(* Logix 5000 project; controller _GigaDiscovery vendor 1 type 14 code 244 rev 35.11; software revision 35.03; part 19 of 23 *)
(* tags used below, declared in another part *)
   CROUT_Air_Compressor : UDT_CROUT;   // Compressor Command -Q18101E
   I_Platform_Closed : UDT_DCM;   // Platform Closed RFID Series -B22501J... -B22807J -B22801B
   I_Platform_Opened : UDT_DCM;   // Platform Opened RFID Series -Q23801J -Q23807J
   No_Sfty : Std_to_Sfty;
   O_Close_Platform : BOOL;
   O_Compressor_Cmd : BOOL;
   O_Open_Platform : BOOL;
   O_Pilots_Valve_Platform : BOOL;
   O_Platform_Main_Valve : BOOL;   // Valvola principale piattaforma B21902I
   O_Platform_MainValve : UDT_CROUT;   // Platform main valve B21902I
   Platform_CloseMain_Valve_Aux_Comand : BOOL;   // Valvola principale piattaforma QV6515E
   Platform_Fbk_Valv_Close : BOOL;   // Platform Close Main Valve Limit Switch -B21909I
   Platform_Fbk_Valv_Open : BOOL;   // Platform Open Main Valve Limit Switch -B21905I
   Platform_OpenMain_Valve_Aux_Comand : BOOL;   // Valvola principale piattaforma QV6515E
   Reset_Pulse : BOOL;
   RESTRAINTS_Rack : LapBar_Racks[41];
   RESTRAINTS_Sector : LapBars_Sector[9];
   Valve_Proof_Test_Cycle : Sequencer;
   Valves_Pressure_Discrepancy : DINT;
(* S_Output, continued *)

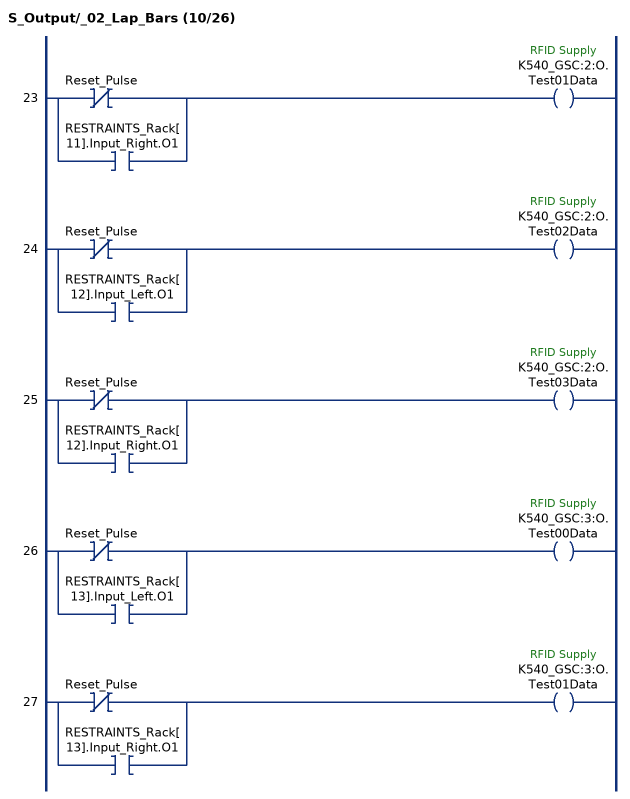
   [picture p369: S_Output/_02_Lap_Bars rungs 23-27]
   23: [XIO(Reset_Pulse) ,XIC(RESTRAINTS_Rack[11].Input_Right.O1) ]OTE(K540_GSC:2:O.Test01Data);
   24: [XIO(Reset_Pulse) ,XIC(RESTRAINTS_Rack[12].Input_Left.O1) ]OTE(K540_GSC:2:O.Test02Data);
   25: [XIO(Reset_Pulse) ,XIC(RESTRAINTS_Rack[12].Input_Right.O1) ]OTE(K540_GSC:2:O.Test03Data);
   26: [XIO(Reset_Pulse) ,XIC(RESTRAINTS_Rack[13].Input_Left.O1) ]OTE(K540_GSC:3:O.Test00Data);
   27: [XIO(Reset_Pulse) ,XIC(RESTRAINTS_Rack[13].Input_Right.O1) ]OTE(K540_GSC:3:O.Test01Data);
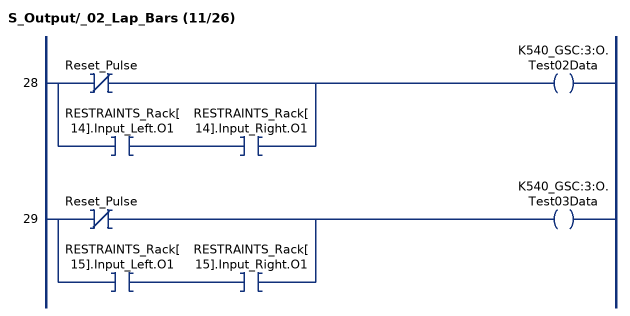
   28: [XIO(Reset_Pulse) ,XIC(RESTRAINTS_Rack[14].Input_Left.O1) XIC(RESTRAINTS_Rack[14].Input_Right.O1) ]OTE(K540_GSC:3:O.Test02Data);
   29: [XIO(Reset_Pulse) ,XIC(RESTRAINTS_Rack[15].Input_Left.O1) XIC(RESTRAINTS_Rack[15].Input_Right.O1) ]OTE(K540_GSC:3:O.Test03Data);
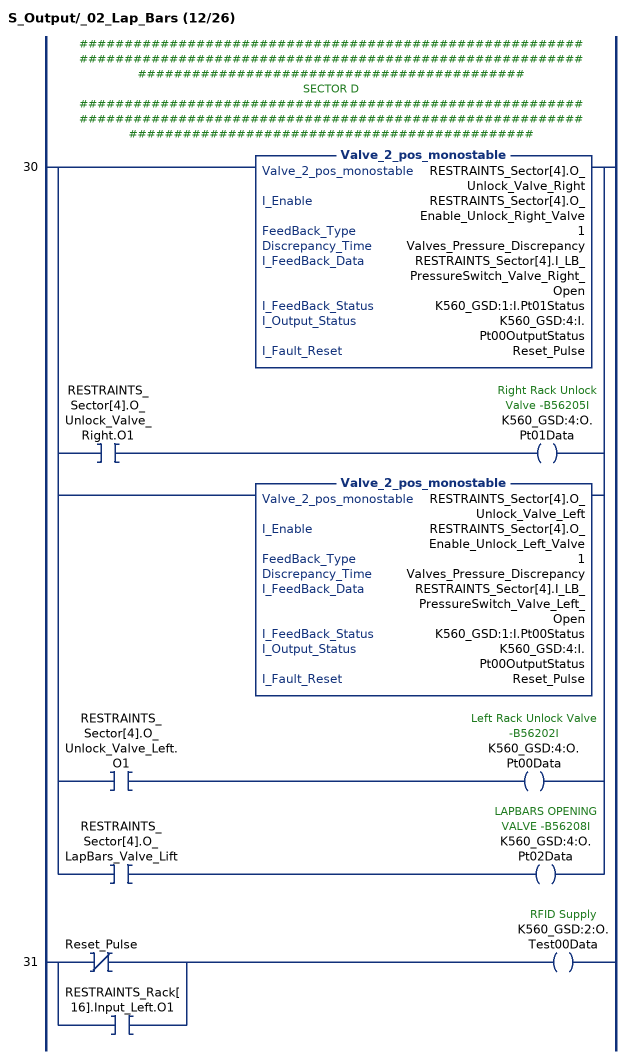
   // ###########################################################################################################################################################
   // SECTOR D
   // #############################################################################################################################################################
   30: [[Valve_2_pos_monostable(RESTRAINTS_Sector[4].O_Unlock_Valve_Right,RESTRAINTS_Sector[4].O_Enable_Unlock_Right_Valve,1,Valves_Pressure_Discrepancy,RESTRAINTS_Sector[4].I_LB_PressureSwitch_Valve_Right_Open,K560_GSD:1:I.Pt01Status,K560_GSD:4:I.Pt00OutputStatus,Reset_Pulse) ,XIC(RESTRAINTS_Sector[4].O_Unlock_Valve_Right.O1) OTE(K560_GSD:4:O.Pt01Data) ] ,[Valve_2_pos_monostable(RESTRAINTS_Sector[4].O_Unlock_Valve_Left,RESTRAINTS_Sector[4].O_Enable_Unlock_Left_Valve,1,Valves_Pressure_Discrepancy,RESTRAINTS_Sector[4].I_LB_PressureSwitch_Valve_Left_Open,K560_GSD:1:I.Pt00Status,K560_GSD:4:I.Pt00OutputStatus,Reset_Pulse) ,XIC(RESTRAINTS_Sector[4].O_Unlock_Valve_Left.O1) OTE(K560_GSD:4:O.Pt00Data) ] ,XIC(RESTRAINTS_Sector[4].O_LapBars_Valve_Lift) OTE(K560_GSD:4:O.Pt02Data) ];
   31: [XIO(Reset_Pulse) ,XIC(RESTRAINTS_Rack[16].Input_Left.O1) ]OTE(K560_GSD:2:O.Test00Data);
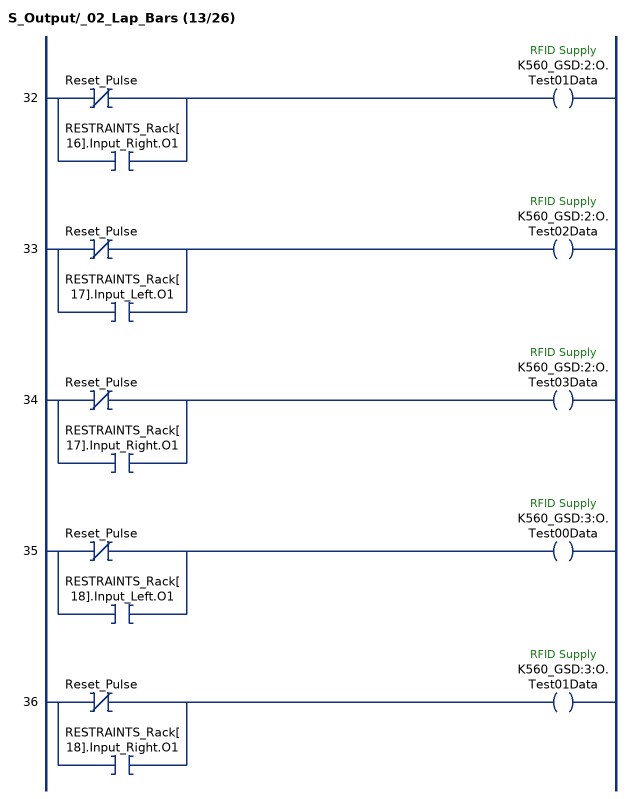
   32: [XIO(Reset_Pulse) ,XIC(RESTRAINTS_Rack[16].Input_Right.O1) ]OTE(K560_GSD:2:O.Test01Data);
   33: [XIO(Reset_Pulse) ,XIC(RESTRAINTS_Rack[17].Input_Left.O1) ]OTE(K560_GSD:2:O.Test02Data);
   34: [XIO(Reset_Pulse) ,XIC(RESTRAINTS_Rack[17].Input_Right.O1) ]OTE(K560_GSD:2:O.Test03Data);
   35: [XIO(Reset_Pulse) ,XIC(RESTRAINTS_Rack[18].Input_Left.O1) ]OTE(K560_GSD:3:O.Test00Data);
   36: [XIO(Reset_Pulse) ,XIC(RESTRAINTS_Rack[18].Input_Right.O1) ]OTE(K560_GSD:3:O.Test01Data);
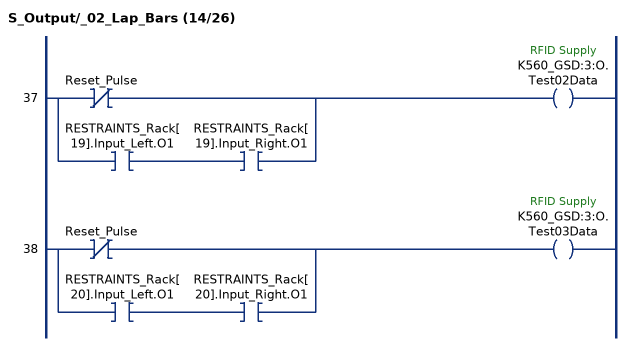
   37: [XIO(Reset_Pulse) ,XIC(RESTRAINTS_Rack[19].Input_Left.O1) XIC(RESTRAINTS_Rack[19].Input_Right.O1) ]OTE(K560_GSD:3:O.Test02Data);
   38: [XIO(Reset_Pulse) ,XIC(RESTRAINTS_Rack[20].Input_Left.O1) XIC(RESTRAINTS_Rack[20].Input_Right.O1) ]OTE(K560_GSD:3:O.Test03Data);
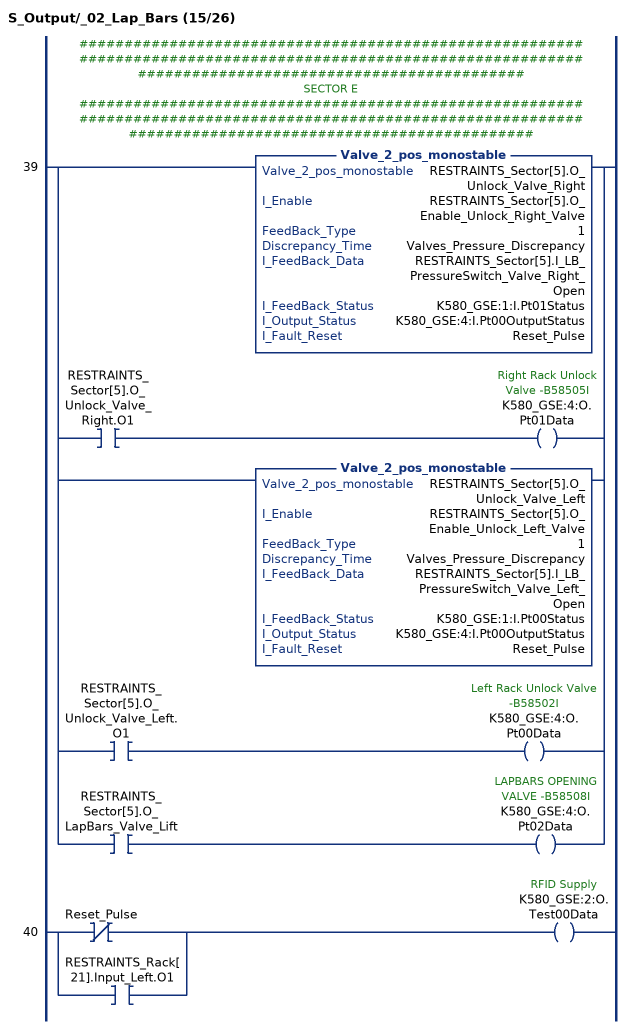
   // ###########################################################################################################################################################
   // SECTOR E
   // #############################################################################################################################################################
   39: [[Valve_2_pos_monostable(RESTRAINTS_Sector[5].O_Unlock_Valve_Right,RESTRAINTS_Sector[5].O_Enable_Unlock_Right_Valve,1,Valves_Pressure_Discrepancy,RESTRAINTS_Sector[5].I_LB_PressureSwitch_Valve_Right_Open,K580_GSE:1:I.Pt01Status,K580_GSE:4:I.Pt00OutputStatus,Reset_Pulse) ,XIC(RESTRAINTS_Sector[5].O_Unlock_Valve_Right.O1) OTE(K580_GSE:4:O.Pt01Data) ] ,[Valve_2_pos_monostable(RESTRAINTS_Sector[5].O_Unlock_Valve_Left,RESTRAINTS_Sector[5].O_Enable_Unlock_Left_Valve,1,Valves_Pressure_Discrepancy,RESTRAINTS_Sector[5].I_LB_PressureSwitch_Valve_Left_Open,K580_GSE:1:I.Pt00Status,K580_GSE:4:I.Pt00OutputStatus,Reset_Pulse) ,XIC(RESTRAINTS_Sector[5].O_Unlock_Valve_Left.O1) OTE(K580_GSE:4:O.Pt00Data) ] ,XIC(RESTRAINTS_Sector[5].O_LapBars_Valve_Lift) OTE(K580_GSE:4:O.Pt02Data) ];
   40: [XIO(Reset_Pulse) ,XIC(RESTRAINTS_Rack[21].Input_Left.O1) ]OTE(K580_GSE:2:O.Test00Data);
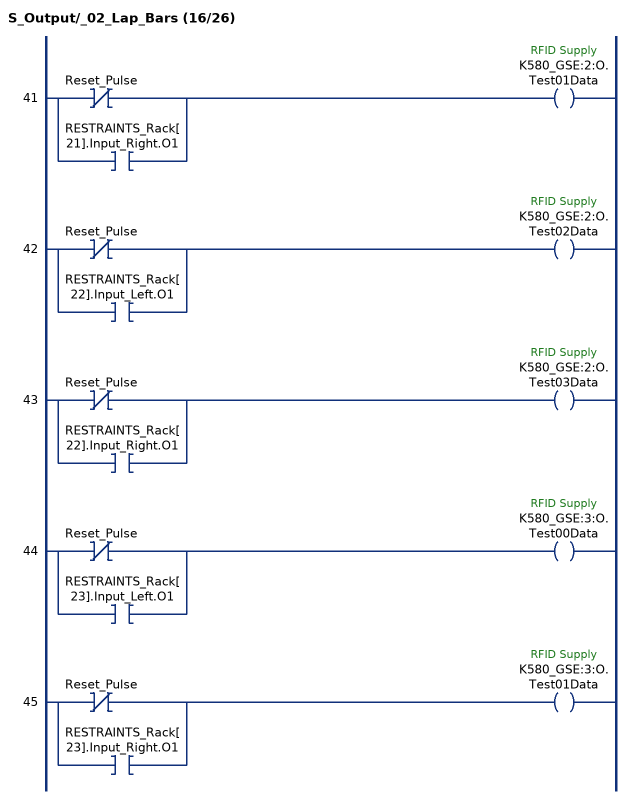
   41: [XIO(Reset_Pulse) ,XIC(RESTRAINTS_Rack[21].Input_Right.O1) ]OTE(K580_GSE:2:O.Test01Data);
   42: [XIO(Reset_Pulse) ,XIC(RESTRAINTS_Rack[22].Input_Left.O1) ]OTE(K580_GSE:2:O.Test02Data);
   43: [XIO(Reset_Pulse) ,XIC(RESTRAINTS_Rack[22].Input_Right.O1) ]OTE(K580_GSE:2:O.Test03Data);
   44: [XIO(Reset_Pulse) ,XIC(RESTRAINTS_Rack[23].Input_Left.O1) ]OTE(K580_GSE:3:O.Test00Data);
   45: [XIO(Reset_Pulse) ,XIC(RESTRAINTS_Rack[23].Input_Right.O1) ]OTE(K580_GSE:3:O.Test01Data);
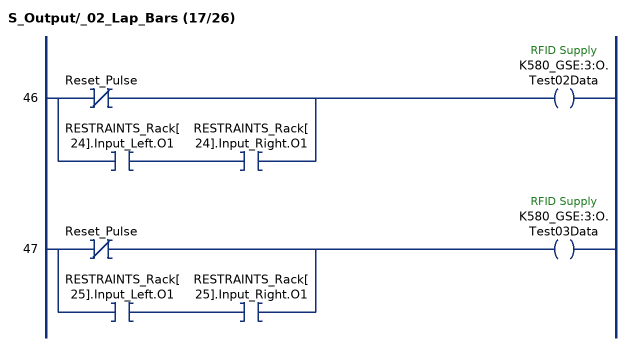
   46: [XIO(Reset_Pulse) ,XIC(RESTRAINTS_Rack[24].Input_Left.O1) XIC(RESTRAINTS_Rack[24].Input_Right.O1) ]OTE(K580_GSE:3:O.Test02Data);
   47: [XIO(Reset_Pulse) ,XIC(RESTRAINTS_Rack[25].Input_Left.O1) XIC(RESTRAINTS_Rack[25].Input_Right.O1) ]OTE(K580_GSE:3:O.Test03Data);
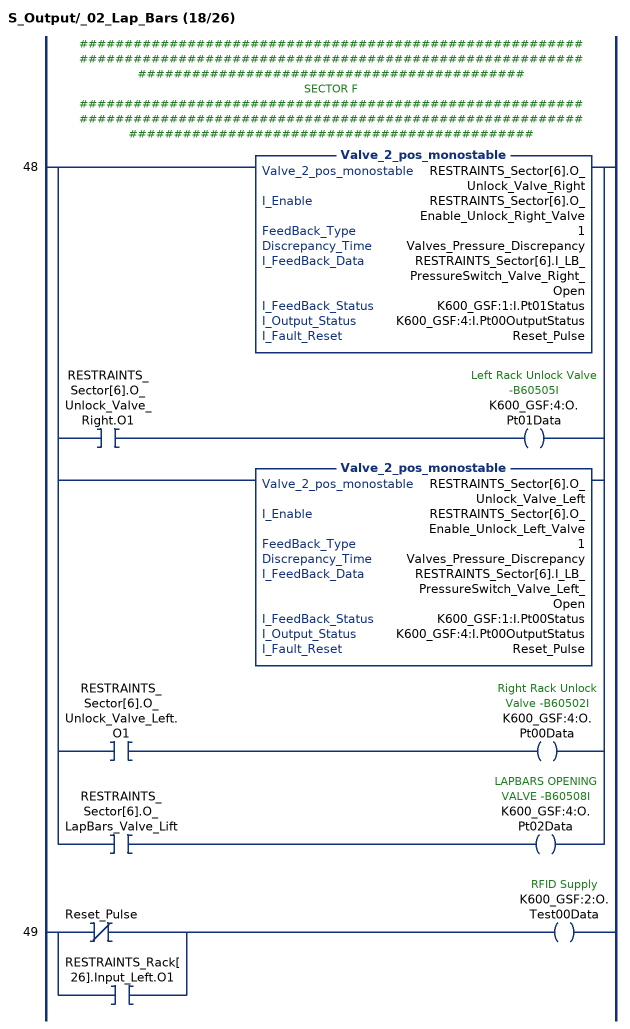
   // ###########################################################################################################################################################
   // SECTOR F
   // #############################################################################################################################################################
   48: [[Valve_2_pos_monostable(RESTRAINTS_Sector[6].O_Unlock_Valve_Right,RESTRAINTS_Sector[6].O_Enable_Unlock_Right_Valve,1,Valves_Pressure_Discrepancy,RESTRAINTS_Sector[6].I_LB_PressureSwitch_Valve_Right_Open,K600_GSF:1:I.Pt01Status,K600_GSF:4:I.Pt00OutputStatus,Reset_Pulse) ,XIC(RESTRAINTS_Sector[6].O_Unlock_Valve_Right.O1) OTE(K600_GSF:4:O.Pt01Data) ] ,[Valve_2_pos_monostable(RESTRAINTS_Sector[6].O_Unlock_Valve_Left,RESTRAINTS_Sector[6].O_Enable_Unlock_Left_Valve,1,Valves_Pressure_Discrepancy,RESTRAINTS_Sector[6].I_LB_PressureSwitch_Valve_Left_Open,K600_GSF:1:I.Pt00Status,K600_GSF:4:I.Pt00OutputStatus,Reset_Pulse) ,XIC(RESTRAINTS_Sector[6].O_Unlock_Valve_Left.O1) OTE(K600_GSF:4:O.Pt00Data) ] ,XIC(RESTRAINTS_Sector[6].O_LapBars_Valve_Lift) OTE(K600_GSF:4:O.Pt02Data) ];
   49: [XIO(Reset_Pulse) ,XIC(RESTRAINTS_Rack[26].Input_Left.O1) ]OTE(K600_GSF:2:O.Test00Data);
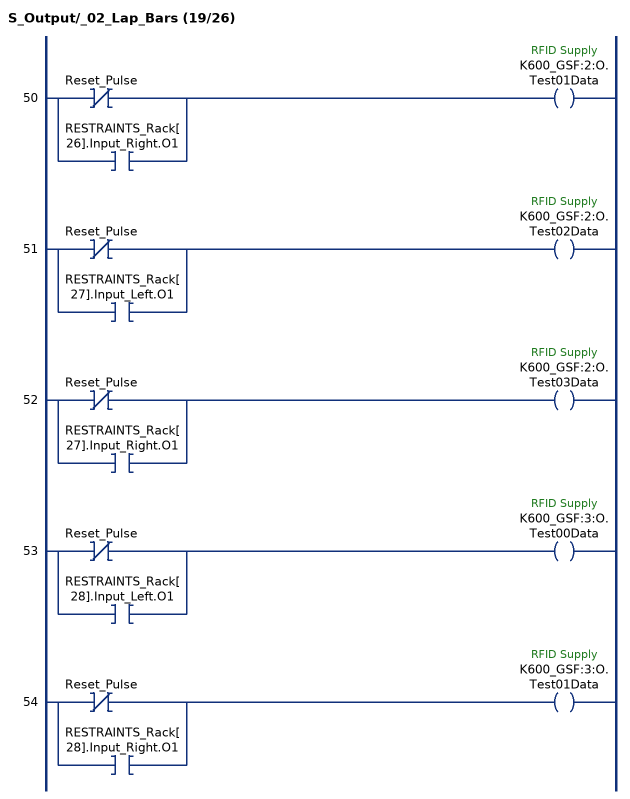
   50: [XIO(Reset_Pulse) ,XIC(RESTRAINTS_Rack[26].Input_Right.O1) ]OTE(K600_GSF:2:O.Test01Data);
   51: [XIO(Reset_Pulse) ,XIC(RESTRAINTS_Rack[27].Input_Left.O1) ]OTE(K600_GSF:2:O.Test02Data);
   52: [XIO(Reset_Pulse) ,XIC(RESTRAINTS_Rack[27].Input_Right.O1) ]OTE(K600_GSF:2:O.Test03Data);
   53: [XIO(Reset_Pulse) ,XIC(RESTRAINTS_Rack[28].Input_Left.O1) ]OTE(K600_GSF:3:O.Test00Data);
   54: [XIO(Reset_Pulse) ,XIC(RESTRAINTS_Rack[28].Input_Right.O1) ]OTE(K600_GSF:3:O.Test01Data);
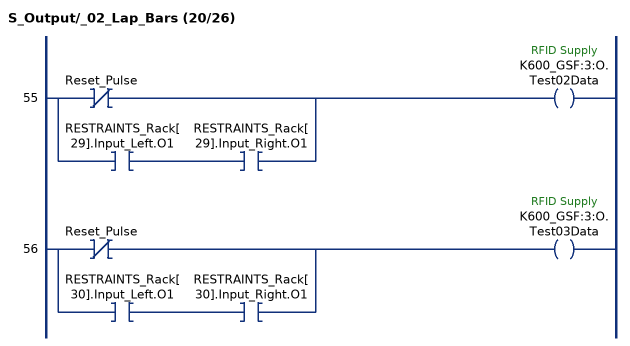
   55: [XIO(Reset_Pulse) ,XIC(RESTRAINTS_Rack[29].Input_Left.O1) XIC(RESTRAINTS_Rack[29].Input_Right.O1) ]OTE(K600_GSF:3:O.Test02Data);
   56: [XIO(Reset_Pulse) ,XIC(RESTRAINTS_Rack[30].Input_Left.O1) XIC(RESTRAINTS_Rack[30].Input_Right.O1) ]OTE(K600_GSF:3:O.Test03Data);
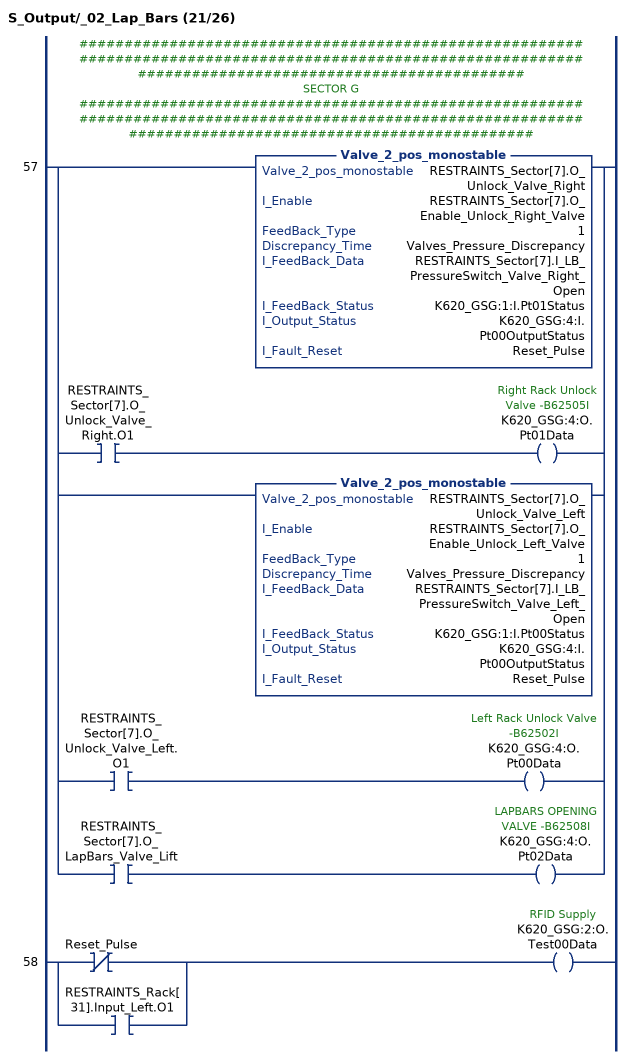
   // ###########################################################################################################################################################
   // SECTOR G
   // #############################################################################################################################################################
   57: [[Valve_2_pos_monostable(RESTRAINTS_Sector[7].O_Unlock_Valve_Right,RESTRAINTS_Sector[7].O_Enable_Unlock_Right_Valve,1,Valves_Pressure_Discrepancy,RESTRAINTS_Sector[7].I_LB_PressureSwitch_Valve_Right_Open,K620_GSG:1:I.Pt01Status,K620_GSG:4:I.Pt00OutputStatus,Reset_Pulse) ,XIC(RESTRAINTS_Sector[7].O_Unlock_Valve_Right.O1) OTE(K620_GSG:4:O.Pt01Data) ] ,[Valve_2_pos_monostable(RESTRAINTS_Sector[7].O_Unlock_Valve_Left,RESTRAINTS_Sector[7].O_Enable_Unlock_Left_Valve,1,Valves_Pressure_Discrepancy,RESTRAINTS_Sector[7].I_LB_PressureSwitch_Valve_Left_Open,K620_GSG:1:I.Pt00Status,K620_GSG:4:I.Pt00OutputStatus,Reset_Pulse) ,XIC(RESTRAINTS_Sector[7].O_Unlock_Valve_Left.O1) OTE(K620_GSG:4:O.Pt00Data) ] ,XIC(RESTRAINTS_Sector[7].O_LapBars_Valve_Lift) OTE(K620_GSG:4:O.Pt02Data) ];
   58: [XIO(Reset_Pulse) ,XIC(RESTRAINTS_Rack[31].Input_Left.O1) ]OTE(K620_GSG:2:O.Test00Data);
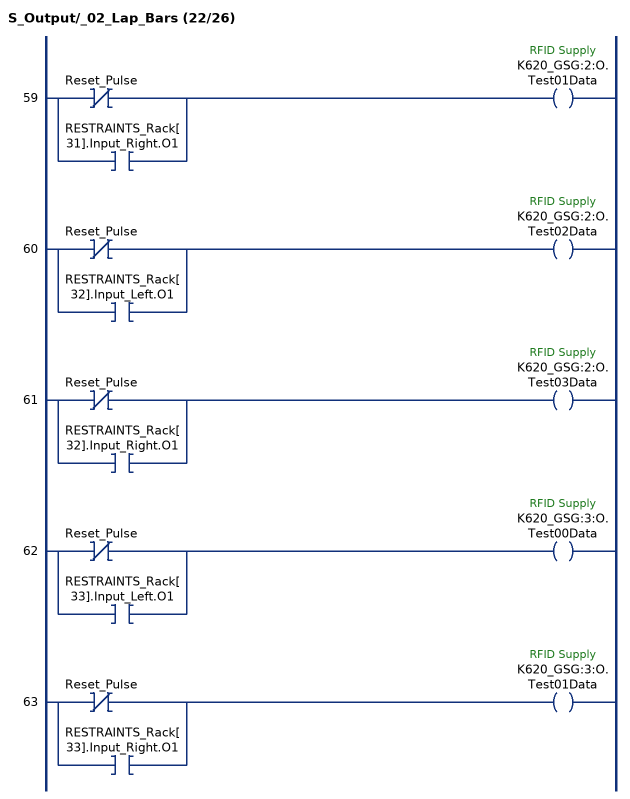
   59: [XIO(Reset_Pulse) ,XIC(RESTRAINTS_Rack[31].Input_Right.O1) ]OTE(K620_GSG:2:O.Test01Data);
   60: [XIO(Reset_Pulse) ,XIC(RESTRAINTS_Rack[32].Input_Left.O1) ]OTE(K620_GSG:2:O.Test02Data);
   61: [XIO(Reset_Pulse) ,XIC(RESTRAINTS_Rack[32].Input_Right.O1) ]OTE(K620_GSG:2:O.Test03Data);
   62: [XIO(Reset_Pulse) ,XIC(RESTRAINTS_Rack[33].Input_Left.O1) ]OTE(K620_GSG:3:O.Test00Data);
   63: [XIO(Reset_Pulse) ,XIC(RESTRAINTS_Rack[33].Input_Right.O1) ]OTE(K620_GSG:3:O.Test01Data);
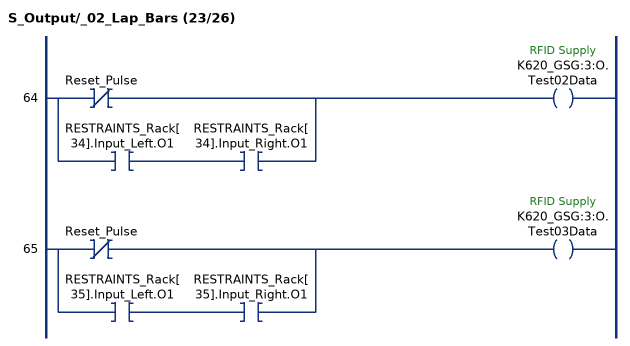
   64: [XIO(Reset_Pulse) ,XIC(RESTRAINTS_Rack[34].Input_Left.O1) XIC(RESTRAINTS_Rack[34].Input_Right.O1) ]OTE(K620_GSG:3:O.Test02Data);
   65: [XIO(Reset_Pulse) ,XIC(RESTRAINTS_Rack[35].Input_Left.O1) XIC(RESTRAINTS_Rack[35].Input_Right.O1) ]OTE(K620_GSG:3:O.Test03Data);
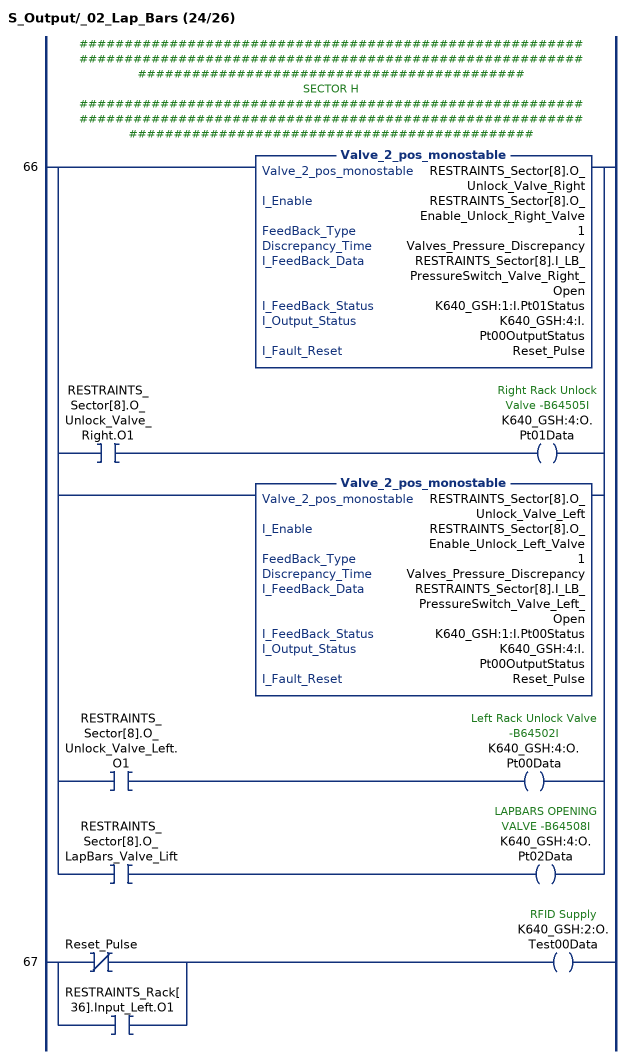
   // ###########################################################################################################################################################
   // SECTOR H
   // #############################################################################################################################################################
   66: [[Valve_2_pos_monostable(RESTRAINTS_Sector[8].O_Unlock_Valve_Right,RESTRAINTS_Sector[8].O_Enable_Unlock_Right_Valve,1,Valves_Pressure_Discrepancy,RESTRAINTS_Sector[8].I_LB_PressureSwitch_Valve_Right_Open,K640_GSH:1:I.Pt01Status,K640_GSH:4:I.Pt00OutputStatus,Reset_Pulse) ,XIC(RESTRAINTS_Sector[8].O_Unlock_Valve_Right.O1) OTE(K640_GSH:4:O.Pt01Data) ] ,[Valve_2_pos_monostable(RESTRAINTS_Sector[8].O_Unlock_Valve_Left,RESTRAINTS_Sector[8].O_Enable_Unlock_Left_Valve,1,Valves_Pressure_Discrepancy,RESTRAINTS_Sector[8].I_LB_PressureSwitch_Valve_Left_Open,K640_GSH:1:I.Pt00Status,K640_GSH:4:I.Pt00OutputStatus,Reset_Pulse) ,XIC(RESTRAINTS_Sector[8].O_Unlock_Valve_Left.O1) OTE(K640_GSH:4:O.Pt00Data) ] ,XIC(RESTRAINTS_Sector[8].O_LapBars_Valve_Lift) OTE(K640_GSH:4:O.Pt02Data) ];
   67: [XIO(Reset_Pulse) ,XIC(RESTRAINTS_Rack[36].Input_Left.O1) ]OTE(K640_GSH:2:O.Test00Data);
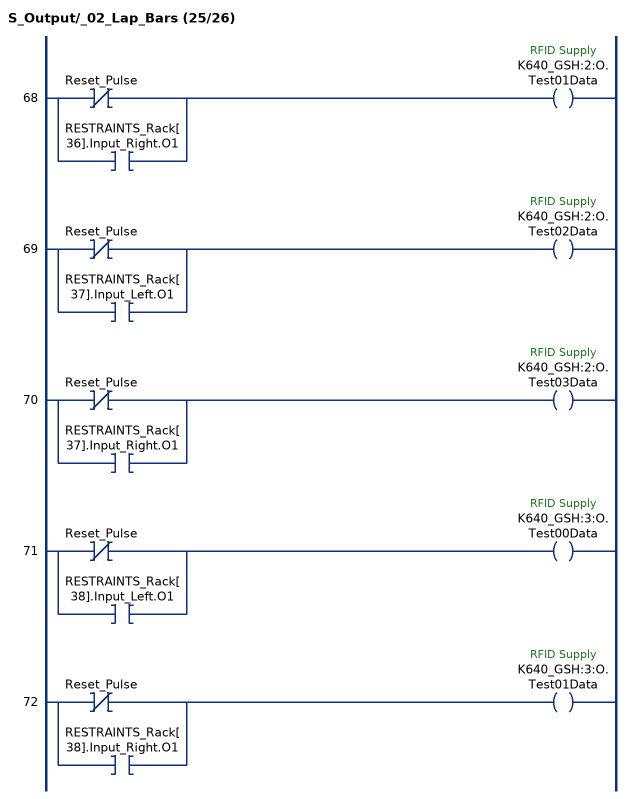
   68: [XIO(Reset_Pulse) ,XIC(RESTRAINTS_Rack[36].Input_Right.O1) ]OTE(K640_GSH:2:O.Test01Data);
   69: [XIO(Reset_Pulse) ,XIC(RESTRAINTS_Rack[37].Input_Left.O1) ]OTE(K640_GSH:2:O.Test02Data);
   70: [XIO(Reset_Pulse) ,XIC(RESTRAINTS_Rack[37].Input_Right.O1) ]OTE(K640_GSH:2:O.Test03Data);
   71: [XIO(Reset_Pulse) ,XIC(RESTRAINTS_Rack[38].Input_Left.O1) ]OTE(K640_GSH:3:O.Test00Data);
   72: [XIO(Reset_Pulse) ,XIC(RESTRAINTS_Rack[38].Input_Right.O1) ]OTE(K640_GSH:3:O.Test01Data);
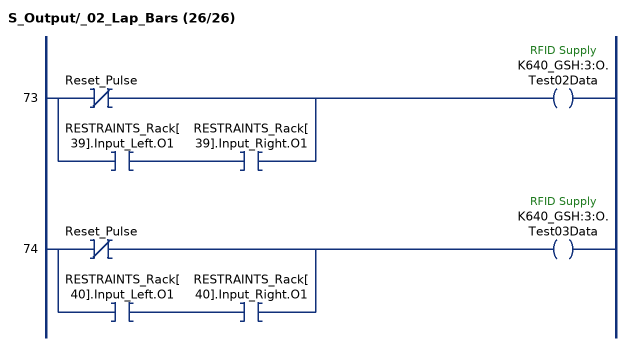
   73: [XIO(Reset_Pulse) ,XIC(RESTRAINTS_Rack[39].Input_Left.O1) XIC(RESTRAINTS_Rack[39].Input_Right.O1) ]OTE(K640_GSH:3:O.Test02Data);
   74: [XIO(Reset_Pulse) ,XIC(RESTRAINTS_Rack[40].Input_Left.O1) XIC(RESTRAINTS_Rack[40].Input_Right.O1) ]OTE(K640_GSH:3:O.Test03Data);
END_ROUTINE

ROUTINE _03_Platform   (* ladder *)
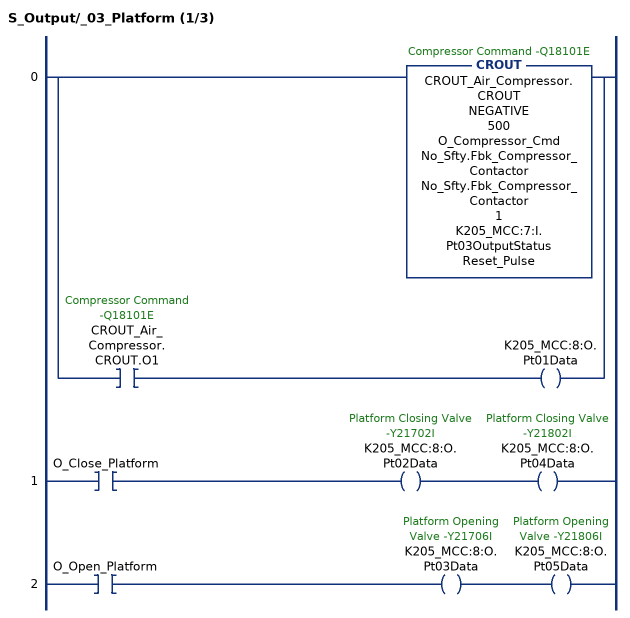
   0: [CROUT(CROUT_Air_Compressor.CROUT,NEGATIVE,500,O_Compressor_Cmd,No_Sfty.Fbk_Compressor_Contactor,No_Sfty.Fbk_Compressor_Contactor,1,K205_MCC:7:I.Pt03OutputStatus,Reset_Pulse) ,XIC(CROUT_Air_Compressor.CROUT.O1) OTE(K205_MCC:8:O.Pt01Data) ];
   1: XIC(O_Close_Platform)OTE(K205_MCC:8:O.Pt02Data)OTE(K205_MCC:8:O.Pt04Data);
   2: XIC(O_Open_Platform)OTE(K205_MCC:8:O.Pt03Data)OTE(K205_MCC:8:O.Pt05Data);
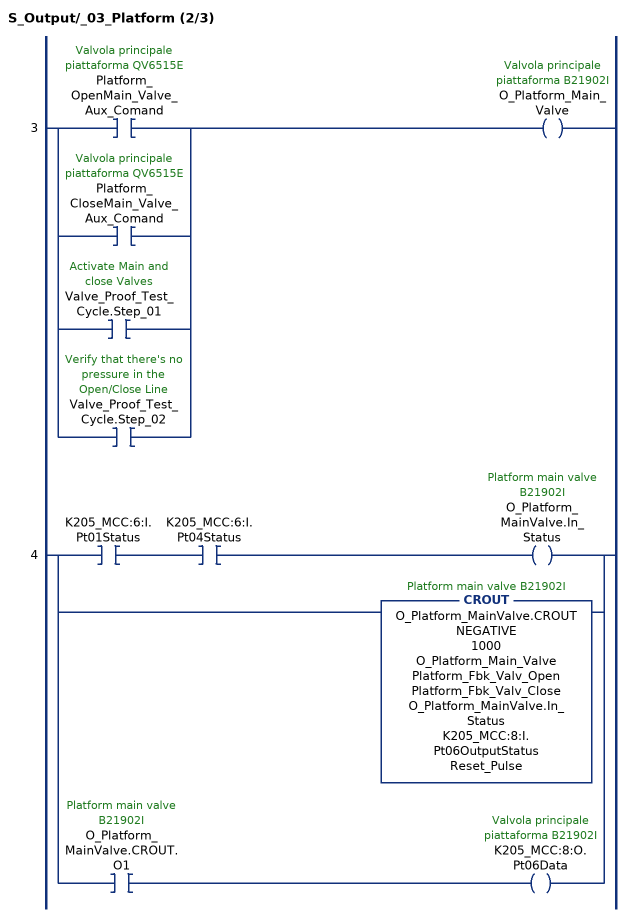
   3: [XIC(Platform_OpenMain_Valve_Aux_Comand) ,XIC(Platform_CloseMain_Valve_Aux_Comand) ,XIC(Valve_Proof_Test_Cycle.Step_01) ,XIC(Valve_Proof_Test_Cycle.Step_02) ]OTE(O_Platform_Main_Valve);
   4: [XIC(K205_MCC:6:I.Pt01Status) XIC(K205_MCC:6:I.Pt04Status) OTE(O_Platform_MainValve.In_Status) ,CROUT(O_Platform_MainValve.CROUT,NEGATIVE,1000,O_Platform_Main_Valve,Platform_Fbk_Valv_Open,Platform_Fbk_Valv_Close,O_Platform_MainValve.In_Status,K205_MCC:8:I.Pt06OutputStatus,Reset_Pulse) ,XIC(O_Platform_MainValve.CROUT.O1) OTE(K205_MCC:8:O.Pt06Data) ];
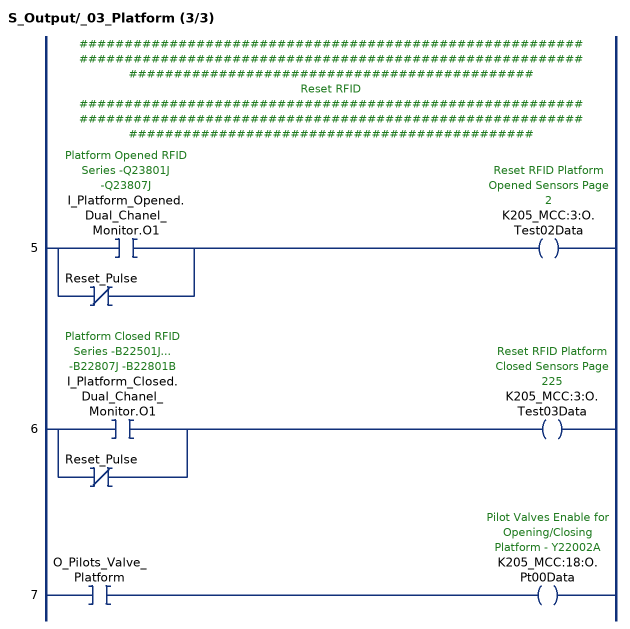
   // #############################################################################################################################################################
   // Reset RFID
   // #############################################################################################################################################################
   5: [XIC(I_Platform_Opened.Dual_Chanel_Monitor.O1) ,XIO(Reset_Pulse) ]OTE(K205_MCC:3:O.Test02Data);
   6: [XIC(I_Platform_Closed.Dual_Chanel_Monitor.O1) ,XIO(Reset_Pulse) ]OTE(K205_MCC:3:O.Test03Data);
   7: XIC(O_Pilots_Valve_Platform)OTE(K205_MCC:18:O.Pt00Data);
END_ROUTINE
